        [0]   // YSV2,FV SYSTEM WORKING BUFFER VESSEL NUMBER
        [2]   // YSV2,TEMPERATURE SETPOINT A. 1/10 DEGREE 'C'
        [30].4   // YSV2,Current vessel final temp.reached
        [4]   // YSV2,TEMPERATURE SETPOINT B. 1/10 DEGREE 'C'
        [6]   // YSV2,TEMPERATURE SETPOINT C. 1/10 DEGREE 'C'
        [8]   // YSV2,TEMPERATURE SETPOINT D. 1/10 DEGREE 'C'
        [36]   // YSV2,Current vessel time to deferred chlling start (hrs.x10)
        [27]   // YSV2,CURRENT ELAPSED HOURS *10
        [40]   // YSV2,FV Routing Status 9=Dirty
        [29]   // YSV2,FLAGS - PLC CONTROL
        [16].1   // YSV2,Profile control flag Hold at B.P B
        [22]   // YSV2,Current FV total residence time
        [16].2   // YSV2,Profile control flag Hold at B.P C
        [29].0   // YSV2,PC TO SAVE TEMPERATURE DATA
        [16].3   // YSV2,Profile control flag Hold at B.P D
        [16].4   // YSV2,Profile control flag Hold at B.P E
        [16].5   // YSV2,Profile control flag Hold at B.P F
        [16].6   // YSV2,Profile control flag Hold at B.P G
        [1]   // YSV2,TEMPERATURE BREAKPOINT A. TIME 1/10 HOURS(ALWAYS=0)
        [29].1   // YSV2,Current vessel deferred chilling enabled flag
        [3]   // YSV2,TEMPERATURE BREAKPOINT B. TIME 1/10 HOURS(ALWAYS=0)
        [5]   // YSV2,TEMPERATURE BREAKPOINT C. TIME 1/10 HOURS(ALWAYS=0)
        [7]   // YSV2,TEMPERATURE BREAKPOINT D. TIME 1/10 HOURS(ALWAYS=0)
        [9]   // YSV2,TEMPERATURE BREAKPOINT E. TIME 1/10 HOURS(ALWAYS=0)
        [11]   // YSV2,TEMPERATURE BREAKPOINT F. TIME 1/10 HOURS(ALWAYS=0)
        [13]   // YSV2,TEMPERATURE BREAKPOINT G. TIME 1/10 HOURS(ALWAYS=0)
        [30].5   // YSV2,Current vessel deferred chilling temp.high flag
        [15].9   // YSV2,Current vessel deferred chilling manual override
   FV_N138 : INT[50] := ([0] := 28, [2] := 30, [3] := 240, [4] := 30, [5] := 480, [6] := 30, [7] := 720, [8] := 30, [9] := 960, [10] := 30, [11] := 1200, [12] := 30, [13] := 32767, [14] := 30, [15] := 20, [17] := -32767, [18] := -32767, [20] := 11748, [22] := 11748, [23] := 1, [25] := 212, [30] := 56);   // YSV3, CURRENT FV DATA
        [15]   // YSV3,FLAGS-PROFILE CONTROL
        [15].4   // YSV3,Profile Control Flags : This is a maturation profile
        [25]   // YSV3,Jacket ACTUAL TEMPERATURE -DEGREES 'C'*10
        [15].5   // YSV3,Profile Control Flags : This is a conditioning profile
        [19]   // YSV3,Current FV max. fermentation time
        [15].2   // YSV3,PLC TO FOLLOW RAMP Breakpoints A to B
        [20]   // YSV3,Current FV warm conditioning time
        [30].3   // YSV3,Current vessel deferred chilling active
        [10]   // YSV3,TEMPERATURE SETPOINT E. 1/10 DEGREE 'C'
        [41]   // YSV3,Cone ACTUAL TEMPERATURE -DEGREES 'C'*10
        [12]   // YSV3,TEMPERATURE SETPOINT F. 1/10 DEGREE 'C'
        [14]   // YSV3,TEMPERATURE SETPOINT G. 1/10 DEGREE 'C'
        [15].3   // YSV3,PLC TO USE CONE COOLING JACKET
        [30].0   // YSV3,Jacket Cooling Valve to open
        [26]   // YSV3,Calculated Setpoint 1/10 degrees C
        [30].1   // YSV3,Cone Cooling Valve to open
        [28]   // YSV3,CURRENT VOLUME HL*10
        [24]   // YSV3,Phase0=No control 1to6 =Fermenting 8 =Pitching Hold 10 =Maturation 11to16=Conditioning
        [0]   // YSV3,FV SYSTEM WORKING BUFFER VESSEL NUMBER
        [2]   // YSV3,TEMPERATURE SETPOINT A. 1/10 DEGREE 'C'
        [30].4   // YSV3,Current vessel final temp.reached
        [4]   // YSV3,TEMPERATURE SETPOINT B. 1/10 DEGREE 'C'
        [6]   // YSV3,TEMPERATURE SETPOINT C. 1/10 DEGREE 'C'
        [8]   // YSV3,TEMPERATURE SETPOINT D. 1/10 DEGREE 'C'
        [36]   // YSV3,Current vessel time to deferred chlling start (hrs.x10)
        [27]   // YSV3,CURRENT ELAPSED HOURS *10
        [40]   // YSV3,FV Routing Status 9=Dirty
        [22]   // YSV3,Current FV total residence time
        [29].0   // YSV3,PC TO SAVE TEMPERATURE DATA
        [29]   // YSV3,FLAGS - PLC CONTROL
        [16].1   // YSV3,Profile control flag Hold at B.P B
        [16].2   // YSV3,Profile control flag Hold at B.P C
        [16].3   // YSV3,Profile control flag Hold at B.P D
        [16].4   // YSV3,Profile control flag Hold at B.P E
        [16].5   // YSV3,Profile control flag Hold at B.P F
        [16].6   // YSV3,Profile control flag Hold at B.P G
        [11]   // YSV3,TEMPERATURE BREAKPOINT F. TIME 1/10 HOURS(ALWAYS=0)
        [1]   // YSV3,TEMPERATURE BREAKPOINT A. TIME 1/10 HOURS(ALWAYS=0)
        [29].1   // YSV3,Current vessel deferred chilling enabled flag
        [3]   // YSV3,TEMPERATURE BREAKPOINT B. TIME 1/10 HOURS(ALWAYS=0)
        [5]   // YSV3,TEMPERATURE BREAKPOINT C. TIME 1/10 HOURS(ALWAYS=0)
        [7]   // YSV3,TEMPERATURE BREAKPOINT D. TIME 1/10 HOURS(ALWAYS=0)
        [9]   // YSV3,TEMPERATURE BREAKPOINT E. TIME 1/10 HOURS(ALWAYS=0)
        [15].9   // YSV3,Current vessel deferred chilling manual override
        [13]   // YSV3,TEMPERATURE BREAKPOINT G. TIME 1/10 HOURS(ALWAYS=0)
        [30].5   // YSV3,Current vessel deferred chilling temp.high flag
   FV_N139 : INT[255] := ([0] := 95, [1] := -32767, [2] := -32767, [3] := -32767, [4] := -32767, [5] := -32767, [6] := -32767, [7] := -32767, [8] := -32767, [9] := -32767, [10] := -32767, [11] := -32767, [12] := -32767, [13] := 32767, [14] := -32767, [15] := 20, [17] := -32767, [18] := -32767, [19] := -32767, [20] := 12650, [21] := -32767, [22] := 32767, [23] := 3, [25] := 184, [30] := 34);   // YST1
        [30].1   // YST1 low level covered flag
        [30].0   // YST1 cooling required
        [0]   // YST1 attemperation control data
   FV_N14 : INT[255] := ([3] := 123);   // ME>PLC Inter PLC comms traf fic outbound
        [0]   // Node 2 Inputs Temporary Depository
        [1]   // Me>FULLERSMV Vessel number just reseeded
        [4]   // Me>FULLERSCT Vessel number just reseeded
        [2].0   // ME>MVSYSTEM Request to change vessel status to ageing
        [5].0   // ME>CTSYSTEM Request to change vessel status to ageing
   FV_N140 : INT[255] := ([0] := 96, [2] := 30, [3] := 240, [4] := 30, [5] := 480, [6] := 30, [7] := 720, [8] := 30, [9] := 960, [10] := 30, [11] := 1200, [12] := 30, [13] := 32767, [14] := 30, [15] := 20, [17] := -32767, [18] := -32767, [20] := 22, [22] := 22, [23] := 1, [24] := 10, [25] := 97, [26] := 30, [27] := 22, [30] := 35);   // YST2
        [30].1   // YST2 low level covered flag
        [30].0   // YST2 cooling required
        [0]   // YST2 attemperation control data
   FV_N141 : INT[255] := ([0] := 5, [1] := 1, [2] := 518, [5] := 518, [7] := 10000, [29] := 2, [30] := 24);   // YSV1 DATA
        [7]   // YSV1 current density
        [4]   // YSV1 startup dialog lock flags
        [3]   // YSV1 Rouser Mode 0=Auto 1 = Manual On 2 = Manual Off
        [5]   // YSV 1 Current Volume Litres
        [4].1   // YSV1 startup by filling pending
        [4].4   // YSV1 startup by waste yeast pending
        [0]   // YSV1 Current Operation
        [2]   // YSV1 current weight kg*10
        [4].5   // YSV1 startup by reseeding pending
        [4].2   // YSV1 startup by pitching pending
        [4].3   // YSV1 startup by cleaning pending
        [6]   // YSV1 current yeast solids percentage
   FV_N142 : INT[255] := ([0] := 5, [1] := 1, [2] := 1551, [5] := 1551, [7] := 10000, [29] := 2, [30] := 24);   // YSV2 DATA
        [4]   // YSV2 startup dialog lock flags
        [5]   // YSV 2 Current Volume Litres
        [4].1   // YSV2 startup by filling pending
        [4].4   // YSV2 startup by waste yeast pending
        [0]   // YSV2 Current Operation
        [2]   // YSV2 current weight kg*10
        [4].2   // YSV2 startup by pitching pending
        [4].3   // YSV2 startup by cleaning pending
   FV_N143 : INT[255] := ([2] := 1, [5] := 1, [7] := 10000, [29] := 2, [30] := 24);   // YSV3 DATA
        [4]   // YSV3 startup dialog lock flags
        [5]   // YSV 3 Current Volume Litres
        [4].1   // YSV3 startup by filling pending
        [0]   // YSV3 Current Operation
        [4].4   // YSV3 startup by waste yeast pending
        [2]   // YSV3 current weight kg*10
        [4].2   // YSV3 startup by pitching pending
        [4].3   // YSV3 startup by cleaning pending
   FV_N144 : INT[255] := ([29] := 2, [30] := 24);   // YST1 DATA
        [4].1   // YST1 start filling pending
        [3]   // YST1 rouser mode: 0=Auto; 1=Manual On; 2=Manual Off
        [4]   // YST1 startup interlock flags
        [4].3   // YST1 start CIP pending
        [0]   // YST1 current operation
   FV_N145 : INT[255] := ([0] := 5, [1] := 1, [29] := 2, [30] := 24);   // YST2 DATA
        [4].1   // YST2 start filling pending
        [3]   // YST1 rouser mode: 0=Auto; 1=Manual On; 2=Manual Off
        [4]   // YST2 startup interlock flags
        [4].3   // YST2 start CIP pending
        [0]   // YST2 current operation
   FV_N146 : INT[50] := ([0] := 226, [2] := 170, [3] := 100, [4] := 190, [5] := 270, [6] := 190, [7] := 300, [8] := 160, [9] := 530, [10] := 160, [11] := 630, [12] := 60, [13] := 32767, [14] := 60, [15] := 64, [16] := 20, [17] := -32767, [18] := -32767, [19] := 1680, [22] := 13, [23] := 1, [24] := 1, [25] := 170, [26] := 190, [27] := 13, [40] := 2, [41] := 171);   // FV26, CURRENT FV DATA
        [15]   // FV26,FLAGS-PROFILE CONTROL
        [15].4   // FV26,Profile Control Flags : This is a maturation profile
        [25]   // FV26,Jacket ACTUAL TEMPERATURE -DEGREES 'C'*10
        [15].5   // FV26,Profile Control Flags : This is a conditioning profile
        [10]   // FV26,TEMPERATURE SETPOINT E. 1/10 DEGREE 'C'
        [15].2   // FV26,PLC TO FOLLOW RAMP Breakpoints A to B
        [19]   // FV26,Current FV max. fermentation time
        [20]   // FV26,Current FV warm conditioning time
        [12]   // FV26,TEMPERATURE SETPOINT F. 1/10 DEGREE 'C'
        [24]   // FV26,Phase0=No control 1to6 =Fermenting 8 =Pitching Hold 10 =Maturation 11to16=Conditioning
        [30].3   // FV26,Current vessel deferred chilling active
        [14]   // FV26,TEMPERATURE SETPOINT G. 1/10 DEGREE 'C'
        [41]   // FV26,Cone ACTUAL TEMPERATURE -DEGREES 'C'*10
        [15].3   // FV26,PLC TO USE CONE COOLING JACKET
        [26]   // FV26,Calculated Setpoint 1/10 degrees C
        [30].0   // FV26,Jacket Cooling Valve to open
        [30].1   // FV26,Cone Cooling Valve to open
        [28]   // FV26,CURRENT VOLUME HL*10
        [0]   // FV26,FV SYSTEM WORKING BUFFER VESSEL NUMBER
        [2]   // FV26,TEMPERATURE SETPOINT A. 1/10 DEGREE 'C'
        [30].4   // FV26,Current vessel final temp.reached
        [4]   // FV26,TEMPERATURE SETPOINT B. 1/10 DEGREE 'C'
        [6]   // FV26,TEMPERATURE SETPOINT C. 1/10 DEGREE 'C'
        [8]   // FV26,TEMPERATURE SETPOINT D. 1/10 DEGREE 'C'
        [27]   // FV26,CURRENT ELAPSED HOURS *10
        [36]   // FV26,Current vessel time to deferred chlling start (hrs.x10)
        [22]   // FV26,Current FV total residence time
        [40]   // FV26,FV Routing Status 9=Dirty
        [29].0   // FV26,PC TO SAVE TEMPERATURE DATA
        [29]   // FV26,FLAGS - PLC CONTROL
        [16].1   // FV26,Profile control flag Hold at B.P B
        [16].2   // FV26,Profile control flag Hold at B.P C
        [16].3   // FV26,Profile control flag Hold at B.P D
        [16].4   // FV26,Profile control flag Hold at B.P E
        [16].5   // FV26,Profile control flag Hold at B.P F
        [16].6   // FV26,Profile control flag Hold at B.P G
        [1]   // FV26,TEMPERATURE BREAKPOINT A. TIME 1/10 HOURS(ALWAYS=0)
        [29].1   // FV26,Current vessel deferred chilling enabled flag
        [3]   // FV26,TEMPERATURE BREAKPOINT B. TIME 1/10 HOURS(ALWAYS=0)
        [11]   // FV26,TEMPERATURE BREAKPOINT F. TIME 1/10 HOURS(ALWAYS=0)
        [13]   // FV26,TEMPERATURE BREAKPOINT G. TIME 1/10 HOURS(ALWAYS=0)
        [5]   // FV26,TEMPERATURE BREAKPOINT C. TIME 1/10 HOURS(ALWAYS=0)
        [7]   // FV26,TEMPERATURE BREAKPOINT D. TIME 1/10 HOURS(ALWAYS=0)
        [30].5   // FV26,Current vessel deferred chilling temp.high flag
        [9]   // FV26,TEMPERATURE BREAKPOINT E. TIME 1/10 HOURS(ALWAYS=0)
        [15].9   // FV26,Current vessel deferred chilling manual override
   FV_N147 : INT[50] := ([0] := 227, [2] := 170, [3] := 100, [4] := 190, [5] := 257, [6] := 190, [7] := 287, [8] := 160, [9] := 517, [10] := 160, [11] := 617, [12] := 60, [13] := 32767, [14] := 60, [15] := 64, [16] := 16, [17] := -32767, [18] := -32767, [19] := 1680, [22] := 492, [23] := 3, [24] := 4, [25] := 159, [26] := 160, [27] := 492, [40] := 3, [41] := 160);   // FV27, CURRENT FV DATA
        [15]   // FV27,FLAGS-PROFILE CONTROL
        [10]   // FV27,TEMPERATURE SETPOINT E. 1/10 DEGREE 'C'
        [25]   // FV27,Jacket ACTUAL TEMPERATURE -DEGREES 'C'*10
        [15].4   // FV27,Profile Control Flags : This is a maturation profile
        [12]   // FV27,TEMPERATURE SETPOINT F. 1/10 DEGREE 'C'
        [19]   // FV27,Current FV max. fermentation time
        [15].5   // FV27,Profile Control Flags : This is a conditioning profile
        [14]   // FV27,TEMPERATURE SETPOINT G. 1/10 DEGREE 'C'
        [41]   // FV27,Cone ACTUAL TEMPERATURE -DEGREES 'C'*10
        [20]   // FV27,Current FV warm conditioning time
        [15].2   // FV27,PLC TO FOLLOW RAMP Breakpoints A to B
        [24]   // FV27,Phase0=No control 1to6 =Fermenting 8 =Pitching Hold 10 =Maturation 11to16=Conditioning
        [30].3   // FV27,Current vessel deferred chilling active
        [15].3   // FV27,PLC TO USE CONE COOLING JACKET
        [26]   // FV27,Calculated Setpoint 1/10 degrees C
        [30].0   // FV27,Jacket Cooling Valve to open
        [30].1   // FV27,Cone Cooling Valve to open
        [0]   // FV27,FV SYSTEM WORKING BUFFER VESSEL NUMBER
        [28]   // FV27,CURRENT VOLUME HL*10
        [2]   // FV27,TEMPERATURE SETPOINT A. 1/10 DEGREE 'C'
        [30].4   // FV27,Current vessel final temp.reached
        [4]   // FV27,TEMPERATURE SETPOINT B. 1/10 DEGREE 'C'
        [6]   // FV27,TEMPERATURE SETPOINT C. 1/10 DEGREE 'C'
        [8]   // FV27,TEMPERATURE SETPOINT D. 1/10 DEGREE 'C'
        [27]   // FV27,CURRENT ELAPSED HOURS *10
        [40]   // FV27,FV Routing Status 9=Dirty
        [22]   // FV27,Current FV total residence time
        [36]   // FV27,Current vessel time to deferred chlling start (hrs.x10)
        [29].0   // FV27,PC TO SAVE TEMPERATURE DATA
        [16].1   // FV27,Profile control flag Hold at B.P B
        [16].2   // FV27,Profile control flag Hold at B.P C
        [16].3   // FV27,Profile control flag Hold at B.P D
        [29]   // FV27,FLAGS - PLC CONTROL
        [1]   // FV27,TEMPERATURE BREAKPOINT A. TIME 1/10 HOURS(ALWAYS=0)
        [16].4   // FV27,Profile control flag Hold at B.P E
        [16].5   // FV27,Profile control flag Hold at B.P F
        [16].6   // FV27,Profile control flag Hold at B.P G
        [11]   // FV27,TEMPERATURE BREAKPOINT F. TIME 1/10 HOURS(ALWAYS=0)
        [29].1   // FV27,Current vessel deferred chilling enabled flag
        [3]   // FV27,TEMPERATURE BREAKPOINT B. TIME 1/10 HOURS(ALWAYS=0)
        [5]   // FV27,TEMPERATURE BREAKPOINT C. TIME 1/10 HOURS(ALWAYS=0)
        [7]   // FV27,TEMPERATURE BREAKPOINT D. TIME 1/10 HOURS(ALWAYS=0)
        [9]   // FV27,TEMPERATURE BREAKPOINT E. TIME 1/10 HOURS(ALWAYS=0)
        [13]   // FV27,TEMPERATURE BREAKPOINT G. TIME 1/10 HOURS(ALWAYS=0)
        [30].5   // FV27,Current vessel deferred chilling temp.high flag
        [15].9   // FV27,Current vessel deferred chilling manual override
   FV_N148 : INT[50] := ([0] := 228, [2] := 170, [3] := 100, [4] := 200, [5] := 290, [6] := 200, [7] := 330, [8] := 200, [9] := 365, [10] := 200, [11] := 475, [12] := 40, [13] := 32767, [14] := 40, [15] := 64, [17] := -32767, [18] := -32767, [19] := 1680, [22] := 1192, [23] := 3, [24] := 6, [25] := 41, [26] := 40, [27] := 1192, [29] := 2, [30] := 24, [40] := 3, [41] := 42);   // FV28, CURRENT FV DATA
        [15]   // FV28,FLAGS-PROFILE CONTROL
        [19]   // FV28,Current FV max. fermentation time
        [10]   // FV28,TEMPERATURE SETPOINT E. 1/10 DEGREE 'C'
        [12]   // FV28,TEMPERATURE SETPOINT F. 1/10 DEGREE 'C'
        [14]   // FV28,TEMPERATURE SETPOINT G. 1/10 DEGREE 'C'
        [41]   // FV28,Cone ACTUAL TEMPERATURE -DEGREES 'C'*10
        [15].4   // FV28,Profile Control Flags : This is a maturation profile
        [25]   // FV28,Jacket ACTUAL TEMPERATURE -DEGREES 'C'*10
        [20]   // FV28,Current FV warm conditioning time
        [15].5   // FV28,Profile Control Flags : This is a conditioning profile
        [15].2   // FV28,PLC TO FOLLOW RAMP Breakpoints A to B
        [24]   // FV28,Phase0=No control 1to6 =Fermenting 8 =Pitching Hold 10 =Maturation 11to16=Conditioning
        [30].3   // FV28,Current vessel deferred chilling active
        [15].3   // FV28,PLC TO USE CONE COOLING JACKET
        [26]   // FV28,Calculated Setpoint 1/10 degrees C
        [30].0   // FV28,Jacket Cooling Valve to open
        [0]   // FV28,FV SYSTEM WORKING BUFFER VESSEL NUMBER
        [2]   // FV28,TEMPERATURE SETPOINT A. 1/10 DEGREE 'C'
        [30].4   // FV28,Current vessel final temp.reached
        [30].1   // FV28,Cone Cooling Valve to open
        [4]   // FV28,TEMPERATURE SETPOINT B. 1/10 DEGREE 'C'
        [6]   // FV28,TEMPERATURE SETPOINT C. 1/10 DEGREE 'C'
        [28]   // FV28,CURRENT VOLUME HL*10
        [8]   // FV28,TEMPERATURE SETPOINT D. 1/10 DEGREE 'C'
        [22]   // FV28,Current FV total residence time
        [27]   // FV28,CURRENT ELAPSED HOURS *10
        [40]   // FV28,FV Routing Status 9=Dirty
        [29].0   // FV28,PC TO SAVE TEMPERATURE DATA
        [36]   // FV28,Current vessel time to deferred chlling start (hrs.x10)
        [1]   // FV28,TEMPERATURE BREAKPOINT A. TIME 1/10 HOURS(ALWAYS=0)
        [29].1   // FV28,Current vessel deferred chilling enabled flag
        [16].1   // FV28,Profile control flag Hold at B.P B
        [16].2   // FV28,Profile control flag Hold at B.P C
        [11]   // FV28,TEMPERATURE BREAKPOINT F. TIME 1/10 HOURS(ALWAYS=0)
        [16].3   // FV28,Profile control flag Hold at B.P D
        [13]   // FV28,TEMPERATURE BREAKPOINT G. TIME 1/10 HOURS(ALWAYS=0)
        [16].4   // FV28,Profile control flag Hold at B.P E
        [16].5   // FV28,Profile control flag Hold at B.P F
        [16].6   // FV28,Profile control flag Hold at B.P G
        [3]   // FV28,TEMPERATURE BREAKPOINT B. TIME 1/10 HOURS(ALWAYS=0)
        [5]   // FV28,TEMPERATURE BREAKPOINT C. TIME 1/10 HOURS(ALWAYS=0)
        [7]   // FV28,TEMPERATURE BREAKPOINT D. TIME 1/10 HOURS(ALWAYS=0)
        [9]   // FV28,TEMPERATURE BREAKPOINT E. TIME 1/10 HOURS(ALWAYS=0)
        [29]   // FV28,FLAGS - PLC CONTROL
        [30].5   // FV28,Current vessel deferred chilling temp.high flag
        [15].9   // FV28,Current vessel deferred chilling manual override
   FV_N149 : INT[50] := ([0] := 229, [2] := 170, [3] := 100, [4] := 190, [5] := 244, [6] := 190, [7] := 274, [8] := 160, [9] := 440, [10] := 160, [11] := 540, [12] := 60, [13] := 32767, [14] := 60, [15] := 64, [17] := -32767, [18] := -32767, [19] := 1680, [22] := 1659, [23] := 3, [25] := 192, [30] := 32, [40] := 9, [41] := 191);   // FV29, CURRENT FV DATA
        [15]   // FV29,FLAGS-PROFILE CONTROL
        [19]   // FV29,Current FV max. fermentation time
        [20]   // FV29,Current FV warm conditioning time
        [10]   // FV29,TEMPERATURE SETPOINT E. 1/10 DEGREE 'C'
        [12]   // FV29,TEMPERATURE SETPOINT F. 1/10 DEGREE 'C'
        [14]   // FV29,TEMPERATURE SETPOINT G. 1/10 DEGREE 'C'
        [41]   // FV29,Cone ACTUAL TEMPERATURE -DEGREES 'C'*10
        [25]   // FV29,Jacket ACTUAL TEMPERATURE -DEGREES 'C'*10
        [15].4   // FV29,Profile Control Flags : This is a maturation profile
        [15].5   // FV29,Profile Control Flags : This is a conditioning profile
        [24]   // FV29,Phase0=No control 1to6 =Fermenting 8 =Pitching Hold 10 =Maturation 11to16=Conditioning
        [30].3   // FV29,Current vessel deferred chilling active
        [15].2   // FV29,PLC TO FOLLOW RAMP Breakpoints A to B
        [15].3   // FV29,PLC TO USE CONE COOLING JACKET
        [26]   // FV29,Calculated Setpoint 1/10 degrees C
        [30].0   // FV29,Jacket Cooling Valve to open
        [0]   // FV29,FV SYSTEM WORKING BUFFER VESSEL NUMBER
        [2]   // FV29,TEMPERATURE SETPOINT A. 1/10 DEGREE 'C'
        [30].4   // FV29,Current vessel final temp.reached
        [4]   // FV29,TEMPERATURE SETPOINT B. 1/10 DEGREE 'C'
        [6]   // FV29,TEMPERATURE SETPOINT C. 1/10 DEGREE 'C'
        [8]   // FV29,TEMPERATURE SETPOINT D. 1/10 DEGREE 'C'
        [30].1   // FV29,Cone Cooling Valve to open
        [28]   // FV29,CURRENT VOLUME HL*10
        [22]   // FV29,Current FV total residence time
        [36]   // FV29,Current vessel time to deferred chlling start (hrs.x10)
        [29].0   // FV29,PC TO SAVE TEMPERATURE DATA
        [27]   // FV29,CURRENT ELAPSED HOURS *10
        [40]   // FV29,FV Routing Status 9=Dirty
        [1]   // FV29,TEMPERATURE BREAKPOINT A. TIME 1/10 HOURS(ALWAYS=0)
        [29].1   // FV29,Current vessel deferred chilling enabled flag
        [3]   // FV29,TEMPERATURE BREAKPOINT B. TIME 1/10 HOURS(ALWAYS=0)
        [11]   // FV29,TEMPERATURE BREAKPOINT F. TIME 1/10 HOURS(ALWAYS=0)
        [16].1   // FV29,Profile control flag Hold at B.P B
        [5]   // FV29,TEMPERATURE BREAKPOINT C. TIME 1/10 HOURS(ALWAYS=0)
        [16].2   // FV29,Profile control flag Hold at B.P C
        [16].3   // FV29,Profile control flag Hold at B.P D
        [16].4   // FV29,Profile control flag Hold at B.P E
        [16].5   // FV29,Profile control flag Hold at B.P F
        [7]   // FV29,TEMPERATURE BREAKPOINT D. TIME 1/10 HOURS(ALWAYS=0)
        [13]   // FV29,TEMPERATURE BREAKPOINT G. TIME 1/10 HOURS(ALWAYS=0)
        [16].6   // FV29,Profile control flag Hold at B.P G
        [9]   // FV29,TEMPERATURE BREAKPOINT E. TIME 1/10 HOURS(ALWAYS=0)
        [30].5   // FV29,Current vessel deferred chilling temp.high flag
        [29]   // FV29,FLAGS - PLC CONTROL
        [15].9   // FV29,Current vessel deferred chilling manual override
   FV_N15 : INT[255] := ([2] := 16, [3] := 14, [4] := 137, [8] := 23, [14] := 14641, [15] := 11826, [16] := 13873, [17] := 11832, [18] := 12338, [19] := 13102, [20] := 50, [64] := 4312, [66] := 16, [67] := 14, [68] := 137, [72] := 23, [78] := 14641, [79] := 11826, [80] := 13873, [81] := 11832, [82] := 12338, [83] := 13102, [84] := 51);   // COMMS_CTRL Inter PLC comms inte rnal working regs
        [63].0   // Status change acknowledgement processing oneshot
        [4].0   // WHT_HL Well Header Tank High Level Probe 0=covered Node 6 Input 0
        [63].1   // Status change acknowledgement processing oneshot
        [0]   // Node 2 Digital Input Word 0
   FV_N150 : INT[50] := ([0] := 230, [2] := 170, [3] := 130, [4] := 190, [5] := 357, [6] := 190, [7] := 437, [8] := 160, [9] := 601, [10] := 160, [11] := 721, [12] := 60, [13] := 32767, [14] := 60, [15] := 64, [17] := -32767, [18] := -32767, [19] := 1680, [20] := 215, [22] := 1895, [23] := 3, [25] := 198, [30] := 32, [40] := 9, [41] := 194);   // FV30, CURRENT FV DATA
        [15]   // FV30,FLAGS-PROFILE CONTROL
        [19]   // FV30,Current FV max. fermentation time
        [20]   // FV30,Current FV warm conditioning time
        [10]   // FV30,TEMPERATURE SETPOINT E. 1/10 DEGREE 'C'
        [12]   // FV30,TEMPERATURE SETPOINT F. 1/10 DEGREE 'C'
        [14]   // FV30,TEMPERATURE SETPOINT G. 1/10 DEGREE 'C'
        [41]   // FV30,Cone ACTUAL TEMPERATURE -DEGREES 'C'*10
        [25]   // FV30,Jacket ACTUAL TEMPERATURE -DEGREES 'C'*10
        [15].4   // FV30,Profile Control Flags : This is a maturation profile
        [15].5   // FV30,Profile Control Flags : This is a conditioning profile
        [24]   // FV30,Phase0=No control 1to6 =Fermenting 8 =Pitching Hold 10 =Maturation 11to16=Conditioning
        [15].3   // FV30,PLC TO USE CONE COOLING JACKET
        [30].3   // FV30,Current vessel deferred chilling active
        [15].2   // FV30,PLC TO FOLLOW RAMP Breakpoints A to B
        [26]   // FV30,Calculated Setpoint 1/10 degrees C
        [22]   // FV30,Current FV total residence time
        [27]   // FV30,CURRENT ELAPSED HOURS *10
        [29].0   // FV30,PC TO SAVE TEMPERATURE DATA
        [30].0   // FV30,Jacket Cooling Valve to open
        [16].1   // FV30,Profile control flag Hold at B.P B
        [16].2   // FV30,Profile control flag Hold at B.P C
        [16].3   // FV30,Profile control flag Hold at B.P D
        [0]   // FV30,FV SYSTEM WORKING BUFFER VESSEL NUMBER
        [2]   // FV30,TEMPERATURE SETPOINT A. 1/10 DEGREE 'C'
        [30].4   // FV30,Current vessel final temp.reached
        [4]   // FV30,TEMPERATURE SETPOINT B. 1/10 DEGREE 'C'
        [30].1   // FV30,Cone Cooling Valve to open
        [6]   // FV30,TEMPERATURE SETPOINT C. 1/10 DEGREE 'C'
        [8]   // FV30,TEMPERATURE SETPOINT D. 1/10 DEGREE 'C'
        [40]   // FV30,FV Routing Status 9=Dirty
        [36]   // FV30,Current vessel time to deferred chlling start (hrs.x10)
        [28]   // FV30,CURRENT VOLUME HL*10
        [1]   // FV30,TEMPERATURE BREAKPOINT A. TIME 1/10 HOURS(ALWAYS=0)
        [29].1   // FV30,Current vessel deferred chilling enabled flag
        [3]   // FV30,TEMPERATURE BREAKPOINT B. TIME 1/10 HOURS(ALWAYS=0)
        [5]   // FV30,TEMPERATURE BREAKPOINT C. TIME 1/10 HOURS(ALWAYS=0)
        [11]   // FV30,TEMPERATURE BREAKPOINT F. TIME 1/10 HOURS(ALWAYS=0)
        [7]   // FV30,TEMPERATURE BREAKPOINT D. TIME 1/10 HOURS(ALWAYS=0)
        [9]   // FV30,TEMPERATURE BREAKPOINT E. TIME 1/10 HOURS(ALWAYS=0)
        [13]   // FV30,TEMPERATURE BREAKPOINT G. TIME 1/10 HOURS(ALWAYS=0)
        [30].5   // FV30,Current vessel deferred chilling temp.high flag
        [16].4   // FV30,Profile control flag Hold at B.P E
        [16].5   // FV30,Profile control flag Hold at B.P F
        [16].6   // FV30,Profile control flag Hold at B.P G
        [29]   // FV30,FLAGS - PLC CONTROL
        [15].9   // FV30,Current vessel deferred chilling manual override
   FV_N151 : INT[50] := ([0] := 231, [2] := 170, [3] := 100, [4] := 190, [5] := 275, [6] := 190, [7] := 305, [8] := 160, [9] := 486, [10] := 160, [11] := 586, [12] := 60, [13] := 32767, [14] := 60, [15] := 64, [17] := -32767, [18] := -32767, [19] := 1680, [20] := 13, [22] := 1693, [23] := 3, [24] := 6, [25] := 60, [26] := 60, [27] := 1693, [29] := 2, [30] := 24, [40] := 3, [41] := 59);   // FV31, CURRENT FV DATA
        [22]   // FV31,Current FV total residence time
        [15]   // FV31,FLAGS-PROFILE CONTROL
        [19]   // FV31,Current FV max. fermentation time
        [20]   // FV31,Current FV warm conditioning time
        [15].3   // FV31,PLC TO USE CONE COOLING JACKET
        [10]   // FV31,TEMPERATURE SETPOINT E. 1/10 DEGREE 'C'
        [12]   // FV31,TEMPERATURE SETPOINT F. 1/10 DEGREE 'C'
        [14]   // FV31,TEMPERATURE SETPOINT G. 1/10 DEGREE 'C'
        [30].0   // FV31,Jacket Cooling Valve to open
        [41]   // FV31,Cone ACTUAL TEMPERATURE -DEGREES 'C'*10
        [11]   // FV31,TEMPERATURE BREAKPOINT F. TIME 1/10 HOURS(ALWAYS=0)
        [25]   // FV31,Jacket ACTUAL TEMPERATURE -DEGREES 'C'*10
        [26]   // FV31,Calculated Setpoint 1/10 degrees C
        [0]   // FV31,FV SYSTEM WORKING BUFFER VESSEL NUMBER
        [2]   // FV31,TEMPERATURE SETPOINT A. 1/10 DEGREE 'C'
        [24]   // FV31,Phase0=No control 1to6 =Fermenting 8 =Pitching Hold 10 =Maturation 11to16=Conditioning
        [29].0   // FV31,PC TO SAVE TEMPERATURE DATA
        [15].4   // FV31,Profile Control Flags : This is a maturation profile
        [30].3   // FV31,Current vessel deferred chilling active
        [15].5   // FV31,Profile Control Flags : This is a conditioning profile
        [15].2   // FV31,PLC TO FOLLOW RAMP Breakpoints A to B
        [27]   // FV31,CURRENT ELAPSED HOURS *10
        [30].4   // FV31,Current vessel final temp.reached
        [16].1   // FV31,Profile control flag Hold at B.P B
        [40]   // FV31,FV Routing Status 9=Dirty
        [1]   // FV31,TEMPERATURE BREAKPOINT A. TIME 1/10 HOURS(ALWAYS=0)
        [16].2   // FV31,Profile control flag Hold at B.P C
        [16].3   // FV31,Profile control flag Hold at B.P D
        [16].4   // FV31,Profile control flag Hold at B.P E
        [16].5   // FV31,Profile control flag Hold at B.P F
        [4]   // FV31,TEMPERATURE SETPOINT B. 1/10 DEGREE 'C'
        [16].6   // FV31,Profile control flag Hold at B.P G
        [6]   // FV31,TEMPERATURE SETPOINT C. 1/10 DEGREE 'C'
        [29].1   // FV31,Current vessel deferred chilling enabled flag
        [28]   // FV31,CURRENT VOLUME HL*10
        [3]   // FV31,TEMPERATURE BREAKPOINT B. TIME 1/10 HOURS(ALWAYS=0)
        [8]   // FV31,TEMPERATURE SETPOINT D. 1/10 DEGREE 'C'
        [5]   // FV31,TEMPERATURE BREAKPOINT C. TIME 1/10 HOURS(ALWAYS=0)
        [7]   // FV31,TEMPERATURE BREAKPOINT D. TIME 1/10 HOURS(ALWAYS=0)
        [30].1   // FV31,Cone Cooling Valve to open
        [13]   // FV31,TEMPERATURE BREAKPOINT G. TIME 1/10 HOURS(ALWAYS=0)
        [9]   // FV31,TEMPERATURE BREAKPOINT E. TIME 1/10 HOURS(ALWAYS=0)
        [36]   // FV31,Current vessel time to deferred chlling start (hrs.x10)
        [30].5   // FV31,Current vessel deferred chilling temp.high flag
        [15].9   // FV31,Current vessel deferred chilling manual override
        [29]   // FV31,FLAGS - PLC CONTROL
   FV_N15_63_0_OutputBit : BOOL;
   FV_N15_63_1_OutputBit : BOOL;
   FV_N16 : INT[255];   // COMMS_TMR Timers used by PLC c omms logic
        [0]   // Node 2 Analogue Input 0 Scaled Value
   FV_N190 : INT[255] := ([2] := 1, [3] := 27, [4] := 1, [102] := 1, [103] := 27, [200] := 8194, [201] := -16384, [203] := 20, [204] := 10, [205] := 137, [206] := 100, [209] := 23, [215] := 14641, [216] := 11826, [217] := 13873, [218] := 11832, [219] := 12338, [220] := 13102, [221] := 52);   // MVR COMMS
        [201]   // Comms to MV Routing PLC
        [200].1   // Enable Comms to MV Routing PLC
   FV_N191 : INT[255] := ([1] := 2, [2] := 3, [3] := 3, [4] := 9, [5] := 9, [6] := 3, [101] := 1, [102] := 4, [103] := 6, [106] := 6, [200] := 2, [201] := -16384, [203] := 20, [204] := 10, [205] := 137, [206] := 100, [209] := 23, [215] := 14641, [216] := 11826, [217] := 13873, [218] := 11832, [219] := 12338, [220] := 13102, [221] := 53);   // FVR COMMS
        [201]   // Comms to FV Routing PLC
        [101]   // FV26Phase0=NoControl 1to6 =Fermenting 8 =Pitching Hold 10 =Maturation 11to16=Conditioning
        [102]   // FV27Phase0=NoControl 1to6 =Fermenting 8 =Pitching Hold 10 =Maturation 11to16=Conditioning
        [103]   // FV28Phase0=NoControl 1to6 =Fermenting 8 =Pitching Hold 10 =Maturation 11to16=Conditioning
        [104]   // FV29Phase0=NoControl 1to6 =Fermenting 8 =Pitching Hold 10 =Maturation 11to16=Conditioning
        [105]   // FV30Phase0=NoControl 1to6 =Fermenting 8 =Pitching Hold 10 =Maturation 11to16=Conditioning
        [200].1   // Enable Comms to FV Routing PLC
        [106]   // FV31Phase0=NoControl 1to6 =Fermenting 8 =Pitching Hold 10 =Maturation 11to16=Conditioning
   FV_N20 : INT[255] := ([1] := -32768, [2] := -32768, [3] := -32768, [4] := -32768, [5] := -32768, [6] := -32768, [7] := -32768);   // YSVFILL<PC YSV Filling data fro m PC
        [0].15   // YSM Filling Startup Cancel Selected
        [0]   // YSV Filling Selected Command
        [1]   // PC>PLC YSV Filling Selected YSV number
        [0].1   // PLC>PC YSM Filling Start Button Selected
        [0].4   // PLC>PC YSV Filling Abort Button Selected
        [0].0   // PC>PLC YSV Filling Startup Dialog Buttlon Selected
        [0].3   // PLC>PC YSV Filling Continue Button Selected
        [0].5   // PLC>PC YSV Filling End Button Selected
        [0].2   // PLC>PC YSV Filling Stop Button Selected
   FV_N21 : INT[255] := ([0] := 1, [2] := 1, [16] := 1, [31] := 3237);   // YSVFILL>PC YSV Filling process data to PC and contr ol regs
        [2]   // YSV Filling Available Commands
        [14]   // YSV Filling Pointer to YSV's Attemporation Data
        [2].3   // PLC>PC YSV Filling Continue Button Available
        [5]   // PLC>PC YSV Filling Process Alarm Parameter (1)
        [9]   // PLC>PC YSV Filling Current Step for PC Display
        [2].2   // PLC>PC YSV Filling Stop Button Available
        [4]   // PLC>PC YSV Filling Process Alarm Number
        [2].0   // PLC>PC YSV Filling Startup Dialog Button Available
        [1]   // YSV Filling Current Step
        [3]   // YSV Filling Restart Step
        [2].1   // PLC>PC YSM Filling Start Button Available
        [15]   // YSV Filling Current YSV data file pointer
        [0]   // YSV Filling Status
        [2].4   // PLC>PC YSV Filling Abort Button Available
        [17]   // YSV Filling Initial YSV weight
        [16]   // YSV Filling Command Processor Step Counter
        [2].5   // PLC>PC YSV Filling End Button Available
   FV_N210 : INT[255] := ([3] := 30, [4] := 30);   // GLYCL_PTRS
        [4]   // Check if Cooling is requested
        [2]   // Clear No of Open Cooling Valves Totaliser
        [0]   // Test for vaild Slot No.
        [3]   // Increment ODD cooling valve totaliser
        [1]   // Clear Slot Number Pointer
   FV_N21_4_alarm : ALARM_DIGITAL;
   FV_N21_4_Alarm_Ready : BOOL;
   FV_N21_4_Delayed_Timer2 : TIMER := (PRE := 1000);
   FV_N21_4_Fault_Returned : STRING;
   FV_N21_4_SQL_Done : DINT := -1;
   FV_N225 : INT[255] := ([0] := 5, [52] := 156, [53] := 18768, [54] := 16706, [61] := 18798, [62] := 25705, [63] := 24864, [64] := 20577, [65] := 27749, [66] := 8257, [67] := 27749, [68] := 8258, [69] := 12107, [77] := 2021, [79] := 24408, [81] := 1178, [82] := 1178, [86] := 2, [87] := 224, [88] := 17, [89] := 4, [90] := 10090, [92] := 2210, [93] := 930);   // GEA DATA FV data to GEA PLCs buffer
   FV_N24 : INT[255] := ([0] := 1, [1] := 2, [2] := 2930);   // YSVFILL_SV YSV filling process data save file to PC
        [0]   // PLC>PC YSV Filling Data Save File 'Save Data Trigger'
        [1]   // PLC>PC YSV Filling Data Save File 'Vessel Filled'
        [2]   // PLC>PC YSV Filling Data Save File 'Weight Filled'
   FV_N245 : INT[255];   // CC_WK_AREA Checkword Work Area
        [27]   // Clear No New Faults Counter
        [3]   // Pointer to de-energised input
        [4].15   // Fault Flag In Checkword
        [4].9   // Desired State Flag In Checkword
        [10].0   // Checking Scan Enabled Latch
        [15].0   // Checkword Unused Flag
        [16]   // No Of Loops To Update All Outputs
        [2]   // Pointer to energised input
        [4].13   // Checking Off Flag In Checkword
        [4].8   // Manual Enabled Flag In Checkword
        [4].11   // De-Energised Input Flag In Checkword
        [11]   // Pointer to Checkword
        [4].10   // Energised Input Flag In Checkword
        [29]   // Preset Value To Be Moved To Fault Counter
   FV_N255 : INT[255] := ([1] := 2112, [2] := 2112, [3] := 2112, [4] := 2112, [5] := 2112, [6] := 2112, [7] := 2368, [8] := 2368, [9] := 2112, [10] := 2112, [11] := 2112, [12] := 2112, [13] := 2112, [14] := 2112, [15] := 2112, [16] := 2112, [17] := 2112, [18] := 2112, [19] := 2112, [20] := 2112, [21] := 2112, [22] := 2112, [23] := 1600, [24] := 1600, [25] := 1600, [26] := 1600, [27] := 2112, [28] := 2112, [29] := 2112, [30] := 2112, [31] := 2112, [32] := 2112, [33] := 2112, [34] := 2112, [35] := 2112, [36] := 2112, [37] := 2112, [38] := 2112, [39] := 2112, [40] := 2112, [41] := 2112, [42] := 2112, [43] := 2112, [44] := 2112, [45] := 2112, [46] := 2112, [47] := 2112, [48] := 2112, [49] := 2112, [50] := 2112, [53] := 2112, [54] := 2112, [55] := 2112, [56] := 2112, [57] := 2112, [58] := 1600, [59] := 2112, [60] := 1600, [61] := 2112, [62] := 1600,
        [63] := 1600, [64] := 2112, [65] := 2128, [66] := 2112, [67] := 2112, [68] := 2112, [69] := 2128, [70] := 2112, [71] := 2112, [72] := 2112, [73] := 2112, [74] := 2080, [75] := 2080, [76] := 1568, [77] := 2368, [78] := 1600, [79] := 2112, [80] := 1600, [81] := 2112, [82] := 2112, [83] := 2112, [84] := 2112, [85] := 2112, [86] := 2112, [87] := 2112, [88] := 2112, [89] := 2112, [90] := 2112, [91] := 2112, [92] := 2112);   // Old Checkwords to keep Delphi working in the interim before full changeover.
   FV_N30 : INT[255] := ([1] := -32768, [2] := -32768, [3] := -32768, [4] := -32768, [5] := -32768, [6] := -32768, [7] := -32768);   // PITCH<PC YSV Pitching data fr om PC
        [0]   // YSV Pitching Selected Command
        [0].3   // PLC>PC YSV Pitching Continue Button Selected
        [2]   // PC>PLC YSV Pitching Required Volume
        [0].2   // PLC>PC YSV Pitching Stop Button Selected
        [1]   // PC>PLC YSV Pitching Selected YSV number
        [0].15   // YSM Pitching Startup Cancel Selected
        [0].1   // PLC>PC YSM Pitching Start Button Selected
        [0].4   // PLC>PC YSV Pitching Abort Button Selected
        [0].5   // PLC>PC YSV Pitching End Button Selected
        [0].0   // PC>PLC YSV Pitching Startup Dialog Buttlon Selected
        [3]   // PC>PLC YSV Pitching FV number being pitched
   FV_N31 : INT[255] := ([0] := 1, [2] := 1, [16] := 1, [17] := 1777, [18] := 1907, [19] := 1575, [20] := 68, [21] := 1562);   // PITCH>PC YSV Pitching data at o PC and control reg isters
        [4]   // PLC>PC YSV Pitching Process Alarm Number
        [2]   // YSV Pitching Available Commands
        [19]   // YSV Pitching Pitch Rate Detection Starting Volume
        [17]   // YSV Pitching Initial YSV volume
        [0]   // YSV Pitching Status
        [18]   // YSV Pitching Max Allowed volume in YSV before Alarming
        [20]   // YSV Pitching Pitch Rate Detection Pitch Rate Litre/min
        [13]   // YSV Pitching Pointer to FV attemporation file
        [2].1   // PLC>PC YSM Pitching Start Button Available
        [2].4   // PLC>PC YSV Pitching Abort Button Available
        [10]   // YPV Pitching Current Volume Pitched Litres
        [16]   // YSV Pitching Command Processor Step Counter
        [2].5   // PLC>PC YSV Pitching End Button Available
        [21]   // YSV Pitching Target Stop Volume in YSV
        [12]   // YSV Pitching YSV operation prior to pitching
        [2].2   // PLC>PC YSV Pitching Stop Button Available
        [5]   // PLC>PC YSV Pitching Process Alarm Parameter (1)
        [9]   // PLC>PC YSV Pitching Current Step for PC Display
        [14]   // YSV Pitching Pointer to YSV's Attemporation Data
        [1]   // YSV Pitching Current Step
        [3]   // YSV Pitching Restart Step
        [2].3   // PLC>PC YSV Pitching Continue Button Available
        [15]   // YSV Pitching Current YSV data file pointer
        [2].0   // PLC>PC YSV Pitching Startup Dialog Button Available
   FV_N31_4_alarm : ALARM_DIGITAL;
   FV_N31_4_Alarm_Ready : BOOL;
   FV_N31_4_Delayed_Timer2 : TIMER := (PRE := 1000);
   FV_N31_4_Fault_Returned : STRING;
   FV_N31_4_SQL_Done : DINT := -1;
   FV_N34 : INT[255] := ([0] := 1, [1] := 2, [2] := 220, [3] := 15);   // PITCH_SV YSV pitching data sa ve file to PC
        [1]   // PLC>PC YSV Pitching Data Save File Vessel Pitched'
        [2]   // PLC>PC YSV Pitching Data Save File Volume Pitched'
        [3]   // PLC>PC YSV Pitching Data Save File FV number pitched
        [0]   // PLC>PC YSV Pitching Data Save File 'Save Data Trigger'
   FV_N40 : INT[255] := ([0] := 32, [1] := -32768, [2] := -32768, [3] := -32768, [4] := -32768, [5] := -32768, [6] := -32768, [7] := -32768);   // YSVCIP<PC
        [0].1   // PLC>PC YSM CIP Start Button Selected
        [0].4   // PLC>PC YSV CIP Abort Button Selected
        [0].0   // PC>PLC YSV CIP Startup Dialog Buttlon Selected
        [1]   // PC>PLC YSV CIP Selected YSV number
        [0].5   // PLC>PC YSV CIP End Button Selected
        [0].2   // PLC>PC YSV CIP Stop Button Selected
        [0].15   // YSM CIP Startup Cancel Selected
        [0]   // YSV CIP Selected Command
        [0].3   // PLC>PC YSV CIP Continue Button Selected
   FV_N41 : INT[255] := ([0] := 1, [2] := 1, [16] := 1);   // YSVCIP>PC
        [2].2   // PLC>PC YSV CIP Stop Button Available
        [2].0   // PLC>PC YSV CIP Startup Dialog Button Available
        [17]   // YSV CIP Initial YSV weight
        [0]   // YSV CIP Status
        [1]   // YSV CIP Current Step
        [3]   // YSV CIP Restart Step
        [2]   // YSV CIP Available Commands
        [14]   // YSV CIP Pointer to YSV's Attemporation Data
        [2].3   // PLC>PC YSV CIP Continue Button Available
        [15]   // YSV CIP Current YSV data file pointer
        [16]   // YSV CIP Command Processor Step Counter
        [2].5   // PLC>PC YSV CIP End Button Available
        [2].1   // PLC>PC YSM CIP Start Button Available
        [2].4   // PLC>PC YSV CIP Abort Button Available
        [4]   // PLC>PC YSV CIP Process Alarm Number
        [5]   // PLC>PC YSV CIP Process Alarm Parameter (1)
        [9]   // PLC>PC YSV CIP Current Step for PC Display
   FV_N41_4_alarm : ALARM_DIGITAL;
   FV_N41_4_Alarm_Ready : BOOL;
   FV_N41_4_Delayed_Timer2 : TIMER := (PRE := 1000);
   FV_N41_4_Fault_Returned : STRING;
   FV_N41_4_SQL_Done : DINT := -1;
   FV_N44 : INT[255];   // YSVCIP_SV
        [0]   // PLC>PC YSV CIP Data Save File 'Save Data Trigger'
        [1]   // PLC>PC YSV CIP Data Save File Vessel CIPed'
        [2]   // PLC>PC YSV CIP Data Save File Weight CIPed'
   FV_N50 : INT[255] := ([1] := -32768, [2] := -32768, [3] := -32768, [4] := -32768, [5] := -32768, [6] := -32768, [7] := -32768);   // WASTE<PC
        [0]   // YSV To Waste Selected Command
        [0].3   // PLC>PC YSV To Waste Continue Button Selected
        [0].2   // PLC>PC YSV To Waste Stop Button Selected
        [1]   // PC>PLC YSV To Waste Selected YSV number
        [0].1   // PLC>PC YSM To Waste Start Button Selected
        [0].4   // PLC>PC YSV To Waste Abort Button Selected
        [0].15   // YSM To Waste Startup Cancel Selected
        [0].5   // PLC>PC YSV To Waste End Button Selected
        [0].0   // PC>PLC YSV To Waste Startup Dialog Buttlon Selected
   FV_N51 : INT[255] := ([0] := 1, [2] := 1, [16] := 1, [17] := 836);   // WASTE>PC
        [0]   // YSV To Waste Status
        [4]   // PLC>PC YSV To Waste Process Alarm Number
        [2]   // YSV To Waste Available Commands
        [13]   // YSV to Waste YSV operation prior to waste transfer
        [17]   // YSV To Waste Initial YSV volume
        [2].1   // PLC>PC YSM To Waste Start Button Available
        [2].4   // PLC>PC YSV To Waste Abort Button Available
        [2].2   // PLC>PC YSV To Waste Stop Button Available
        [16]   // YSV To Waste Command Processor Step Counter
        [2].5   // PLC>PC YSV To Waste End Button Available
        [5]   // PLC>PC YSV To Waste Process Alarm Parameter (1)
        [14]   // YSV To Waste Pointer to YSV's Attemporation Data
        [9]   // PLC>PC YSV To Waste Current Step for PC Display
        [1]   // YSV To Waste Current Step
        [2].3   // PLC>PC YSV To Waste Continue Button Available
        [3]   // YSV To Waste Restart Step
        [15]   // YSV To Waste Current YSV data file pointer
        [2].0   // PLC>PC YSV To Waste Startup Dialog Button Available
   FV_N51_4_alarm : ALARM_DIGITAL;
   FV_N51_4_Alarm_Ready : BOOL;
   FV_N51_4_Delayed_Timer2 : TIMER := (PRE := 1000);
   FV_N51_4_Fault_Returned : STRING;
   FV_N51_4_SQL_Done : DINT := -1;
   FV_N54 : INT[255] := ([0] := 1, [1] := 2, [2] := 830);   // WASTE_SV
        [2]   // PLC>PC YSV To Waste Data Save File Volume Transfered
        [3]   // PLC>PC YSV To Waste Data Save File FV number pitched
        [1]   // PLC>PC YSV To Waste Data Save File YSV number
        [0]   // PLC>PC YSV To Waste Data Save File 'Save Data Trigger'
   FV_N60 : INT[255] := ([1] := -32768, [2] := -32768, [3] := -32768, [4] := -32768, [5] := -32768, [6] := -32768, [7] := -32768);   // RESEED<PC
        [3]   // Source Vessel
        [0]   // YSV Reseeding Selected Command
        [0].2   // PLC>PC YSV Reseeding Stop Button Selected
        [0].1   // PLC>PC YSM Reseeding Start Button Selected
        [0].4   // PLC>PC YSV Reseeding Abort Button Selected
        [0].0   // PC>PLC YSV Reseeding Startup Dialog Buttlon Selected
        [0].5   // PLC>PC YSV Reseeding End Button Selected
        [1]   // PC>PLC YSV Reseeding Selected YSV number
        [0].3   // PLC>PC YSV Reseeding Continue Button Selected
        [2]   // Reseeding Volume
        [0].15   // YSM Reseeding Startup Cancel Selected
        [4]   // PC>PLC Reseeding Destination vessel number
   FV_N61 : INT[255] := ([0] := 1, [2] := 1, [16] := 1, [17] := 526, [18] := 656, [21] := 520);   // RESEED>PC
        [17]   // Reseeding initial YSV volume
        [10]   // Reseeding total volume transferred for PC display
        [14]   // YSV Reseeding Pointer to YSV's Attemporation Data
        [2].3   // PLC>PC YSV Reseeding Continue Button Available
        [21]   // Reseeding target end volume
        [5]   // PLC>PC YSV Reseeding Process Alarm Parameter (1)
        [9]   // PLC>PC YSV Reseeding Current Step for PC Display
        [16]   // YSV Reseeding Command Processor Step Counter
        [0]   // YSV Reseeding Status
        [19]   // Reseeding last discharge weight check weight
        [1]   // YSV Reseeding Current Step
        [3]   // YSV Reseeding Restart Step
        [2].5   // PLC>PC YSV Reseeding End Button Available
        [2].2   // PLC>PC YSV Reseeding Stop Button Available
        [2].0   // PLC>PC YSV Reseeding Startup Dialog Button Available
        [15]   // YSV Reseeding Current YSV data file pointer
        [20]   // Reseeding Weight lost in last 60 secs
        [18]   // Reseeding max.vol. allowed before alarm
        [2].1   // PLC>PC YSM Reseeding Start Button Available
        [2].4   // PLC>PC YSV Reseeding Abort Button Available
        [13]   // YSV reseeding pointer to FV's attemperation file
        [4]   // PLC>PC YSV Reseeding Process Alarm Number
        [2]   // YSV Reseeding Available Commands
   FV_N61_4_alarm : ALARM_DIGITAL;
   FV_N61_4_Alarm_Ready : BOOL;
   FV_N61_4_Delayed_Timer2 : TIMER := (PRE := 1000);
   FV_N61_4_Fault_Returned : STRING;
   FV_N61_4_SQL_Done : DINT := -1;
   FV_N64 : INT[255] := ([0] := 1, [1] := 1, [2] := 6, [3] := 7, [4] := 37);   // RESEED_SV
        [2]   // PLC>PC YSV Reseeding Data Save File Volume Reseeded'
        [0].0   // PLC>PC Reseeding save data flag
        [1]   // PLC>PC YSV Reseeding Data Save File YSV number
        [3]   // PLC>PC YSV Reseeding Data Save File FV reseeded
        [4]   // PLC>PC YSV Reseeding Data Save File MV reseeded
        [0]   // PLC>PC YSV Reseeding Data Save File 'Save Data Trigger'
   FV_N7 : INT[255] := ([0] := -42);   // INTEGER
        [0]   // Glycol tank temperature -15.0 to 10.0 C
   FV_N70 : INT[255];   // LNCIP <PC
        [0].0   // PC>PLC Line CIP startup dialog button selected
        [0].5   // PC > PLC Line CIP end selected
        [1]   // PC>PLC Line CIP Selected YSV number
        [0].3   // PC > PLC Line CIP continue button selected
        [0].1   // Line CIP start selected
        [0].2   // PC > PLC Line CIP stop button selected
        [0]   // Line CIP selected command
        [0].4   // PC > PLC Line CIP abort button selected
        [0].15   // Line CIP startup cancelled
   FV_N71 : INT[255] := ([0] := 1, [2] := 1, [16] := 1);   // LNCIP >PC
        [16]   // Line CIP Command Processor Step Counter
        [2].2   // PLC>PC Line CIP stop button available
        [2].0   // PLC>PC Line CIP startup dialog button available
        [0]   // Line CIP status
        [4]   // PLC>PC Reeseeding process Current alarm number
        [2].3   // PLC>PC Line CIP continue button available
        [2].1   // PLC>PC Line CIP start button available
        [2].5   // PLC>PC Line CIP end button available
        [2].4   // PLC>PC Line CIP abort button available
        [5]   // PLC>PC Reseeding process Alarm parameter 1
        [1]   // Line CIP current step
        [3]   // Line CIP restart step
        [9]   // PLC>PC Line CIP current step for PC display
   FV_N71_4_alarm : ALARM_DIGITAL;
   FV_N71_4_Alarm_Ready : BOOL;
   FV_N71_4_Delayed_Timer2 : TIMER := (PRE := 1000);
   FV_N71_4_Fault_Returned : STRING;
   FV_N71_4_SQL_Done : DINT := -1;
   FV_N80 : INT[255] := ([1] := -32768, [2] := -32768, [3] := -32768, [4] := -32768, [5] := -32768, [6] := -32768, [7] := -32768);   // YSTFILL<PC YST filling data fro m PC
        [0].5   // End YST filling
        [0].2   // Stop YST filling
        [0].1   // Start YST filling
        [0].4   // Abort YST filling
        [0]   // YST filling selected command
        [1]   // YST filling selected YST
        [0].3   // Continue YST filling
        [0].0   // Initiate YST filling startup
        [0].15   // YST filling cancel startup
   FV_N81 : INT[255] := ([0] := 1, [2] := 1, [16] := 1);   // YSTFILL>PC YST filling process data to PC and contr ol regs.
        [2].5   // YST filling end available
        [2].2   // YST filling stop available
        [2].1   // YST filling start available
        [2].4   // YST filling abort available
        [0]   // YST filling status (0:Unavailable; 1:Idle; 2:Running; 3:Stopped; 4:Faulted)
        [14]   // YST filling current YST attemperation file pointer
        [2].3   // YST filling continue available
        [4]   // YST filling routine alarm register
        [1]   // YST filling current step
        [2].0   // YST filling initiate startup available
        [3]   // YST filling restart step
        [9]   // YST filling PC- displayed current step
